FUNCTION_BLOCK UConveyor
VAR
  iStep : INT;
END_VAR
VAR_IN_OUT
  ConveyorIOLeft : ConveyorIO;  (* U的左半边 *)
  ConveyorIORight : ConveyorIO;  (* U的右半边 *)
  ConveyorIODown : ConveyorIO;  (* U的下边一横 *)
  UConveyorIO : UConveyorIO;  (* 顶升,阻挡 *)
END_VAR
VAR
  m_xInitial : BOOL;
  m_tonCylinderOvertime : TON;  (* 气缸超时报警定时器 *)
  m_tCylinderOvertimeCurrent : TIME;
  m_tonExitBarDelay : TON;  (* 退出阻挡器延时 *)
  m_tExitBarDelay : TIME;
  m_xExitBarDelay : BOOL;
  m_TonStep0 : TON;  (* Step为0延时 *)
  m_xStep0 : BOOL;  (* Step为0延时 *)
  m_tStep0 : TIME;  (* Step为0延时 *)
END_VAR
(*                                                                                                          
初始化中增加气缸复位，气缸位置有BUG
//*)
IF NOT m_xInitial THEN
	UConveyorIO.tSetOvertime:=T#5s;
	UConveyorIO.xExitEnable1:=1;
	UConveyorIO.xExitEnable2:=1;
	UConveyorIO.xExitEnable3:=1;
	m_xInitial:=1;
END_IF;
(*外部不用写ConveyorDown的开关，会自己根据来料的产品信息判断停哪个光电*)
IF UConveyorIO.iTask=1 AND ConveyorIODown.diDesConveyorIn=ConveyorIOLeft.diDeviceID THEN
	ConveyorIODown.xCWPresent:=ConveyorIOLeft.xCCWPresent;
ELSIF UConveyorIO.iTask=1 AND ConveyorIODown.diDesConveyorIn=ConveyorIORight.diDeviceID THEN
	ConveyorIODown.xCWPresent:=ConveyorIORight.xCCWPresent;
ELSE
	ConveyorIODown.xCWPresent:=ConveyorIOLeft.xCCWPresent OR ConveyorIORight.xCCWPresent;
END_IF;
(*这里判断什么时候直接放行，左右都不需要，也不是0，就放走*)
IF  NOT(ConveyorIODown.diDesConveyor=ConveyorIOLeft.diDeviceID 
		OR  ConveyorIODown.diDesConveyor=ConveyorIORight.diDeviceID 
		OR ConveyorIODown.diDesConveyor=0) THEN
	UConveyorIO.xPassEnable:=1;
ELSE
	UConveyorIO.xPassEnable:=0;
END_IF;	
IF g_xAuto THEN	
(*	//加个Step为0的延时，防止扫描周期的影响*)
	m_TonStep0(IN:= iStep=0 ,PT:= t#100ms ,Q:= m_xStep0 ,ET:= m_tStep0 );
	(*//这个是留给阻挡动作的时间*)
	m_tonExitBarDelay(IN:=iStep=4 ,PT:= T#1s ,Q:= m_xExitBarDelay ,ET:= m_tExitBarDelay);
CASE UConveyorIO.iTask OF(*这个Task做抢占，可做LastTask保护*)
0:(*各种初始化，能自动去3*)
	ConveyorIODown.xLoad:=0;
	ConveyorIOleft.xLoad:=0;
	ConveyorIORight.xLoad:=0;
	ConveyorIODown.xUnload:=0;
	ConveyorIOLeft.xUnload:=0;
	ConveyorIORight.xUnload:=0;
	ConveyorIODown.xPutInto:=0;
	ConveyorIOLeft.xPutInto:=0;
	ConveyorIORight.xPutInto:=0;	
	UConveyorIO.xExitBarCylinderRetract1:=0;
	UConveyorIO.xExitBarCylinderRetract2:=0;	
	UConveyorIO.xLiftCylinderRetract1:=1;
	UConveyorIO.xLiftCylinderRetract2:=1;
	UConveyorIO.xLiftCylinderExtend1:=0;
	UConveyorIO.xLiftCylinderExtend2:=0;
1:(*上料*)
	CASE iStep OF
	0:(*各种初始化，能自动去3*)
		ConveyorIODown.xLoad:=0;
		ConveyorIOleft.xLoad:=0;
		ConveyorIORight.xLoad:=0;
		ConveyorIODown.xUnload:=0;
		ConveyorIOLeft.xUnload:=0;
		ConveyorIORight.xUnload:=0;
		UConveyorIO.xExitBarCylinderRetract1:=0;
		UConveyorIO.xExitBarCylinderRetract2:=0;
		UConveyorIO.xBatteryError:=0;
		ConveyorIODown.xPutInto:=0;
		ConveyorIOLeft.xPutInto:=0;
		ConveyorIORight.xPutInto:=0;	
	(*	//根据是否有料判断去1还是3，但会等一个延时*)
		IF m_xStep0 AND  ConveyorIODown.xEmpty THEN
			iStep:=1;
		ELSIF m_xStep0 AND NOT ConveyorIODown.xEmpty THEN
			iStep:=3;
		END_IF;	
	1:(*顶升初始化，等load*)
		(*//左顶升*)
		IF UConveyorIO.xLiftCylinderExtendInit1 THEN
			UConveyorIO.xLiftCylinderExtend1:=1;
			UConveyorIO.xLiftCylinderRetract1:=0;
		ELSE
			UConveyorIO.xLiftCylinderExtend1:=0;
			UConveyorIO.xLiftCylinderRetract1:=1;
		END_IF;
	(*	//右顶升*)
		IF UConveyorIO.xLiftCylinderExtendInit2 THEN
			UConveyorIO.xLiftCylinderExtend2:=1;
			UConveyorIO.xLiftCylinderRetract2:=0;
			ELSE
			UConveyorIO.xLiftCylinderExtend2:=0;
			UConveyorIO.xLiftCylinderRetract2:=1;
		END_IF;
		(*//顶升到位，等上料信号*)
		IF 	((UConveyorIO.xLiftCylinderExtendInit1 AND UConveyorIO.xLiftCylinderExtendDetect1)
				OR (NOT UConveyorIO.xLiftCylinderExtendInit1 AND UConveyorIO.xLiftCylinderRetractDetect1))
			AND	((UConveyorIO.xLiftCylinderExtendInit2 AND UConveyorIO.xLiftCylinderExtendDetect2)
		   		OR (NOT UConveyorIO.xLiftCylinderExtendInit2 AND UConveyorIO.xLiftCylinderRetractDetect2))		
			AND	UConveyorIO.xEntryEnable1 THEN(*有上料请求1*)
		   	ConveyorIODown.xLoad:=1;
			iStep:=2;
		END_IF;
	2:(*Load完成*)
		(*去右臂时才需要阻挡1放行,其他情况阻挡1挡住*)
		UConveyorIO.xExitBarCylinderRetract1:=ConveyorIODown.diDesConveyorIn=ConveyorIORight.diDeviceID;
		IF NOT ConveyorIODown.xEmpty THEN
			ConveyorIODown.xLoad:=0;
			ConveyorIOLeft.xPutInto:=1;
			ConveyorIOright.xPutInto:=1;
			istep:=3;
		END_IF;
	3:(*顶升等Unload，这里等有了ExitEnable再顶升，因为可能有地方需要允许了再升降，比如倍速链*)
		(*//电池检测保护，防止把带电池的料框送进去了*)
		IF (ConveyorIODown.diDesConveyor=ConveyorIOLeft.diDeviceID OR ConveyorIODown.diDesConveyor=ConveyorIORight.diDeviceID)
			AND	(UConveyorIO.xBatteryDetect1 OR UConveyorIO.xBatteryDetect2)(*在下面时检测*)
			AND UConveyorIO.xLiftCylinderRetractDetect1 AND UConveyorIO.xLiftCylinderRetractDetect2 THEN
			UConveyorIO.xBatteryError:=1;
		END_IF;	
		(*//左侧顶升控制*)
		IF (ConveyorIODown.diDesConveyor=ConveyorIOLeft.diDeviceID AND UConveyorIO.xExitEnable2 AND NOT UConveyorIO.xBatteryError)THEN
			IF UConveyorIO.xLiftCylinderExtendInit1 THEN
				UConveyorIO.xLiftCylinderExtend1:=0;
				UConveyorIO.xLiftCylinderRetract1:=1;
			ELSE
				UConveyorIO.xLiftCylinderExtend1:=1;
				UConveyorIO.xLiftCylinderRetract1:=0;
			END_IF;
			IF(NOT UConveyorIO.xLiftCylinderExtendInit1 AND UConveyorIO.xLiftCylinderExtendDetect1)
				OR (UConveyorIO.xLiftCylinderExtendInit1 AND UConveyorIO.xLiftCylinderRetractDetect1)THEN
				ConveyorIOLeft.xPutInto:=0;
				ConveyorIOright.xPutInto:=0;
				iStep:=4;
			END_IF;
		END_IF;	
		(*//右侧顶升控制*)
		IF (ConveyorIODown.diDesConveyor=ConveyorIORight.diDeviceID AND UConveyorIO.xExitEnable3 AND NOT UConveyorIO.xBatteryError)THEN
			IF UConveyorIO.xLiftCylinderExtendInit2 THEN
				UConveyorIO.xLiftCylinderExtend2:=0;
				UConveyorIO.xLiftCylinderRetract2:=1;
			ELSE
				UConveyorIO.xLiftCylinderExtend2:=1;
				UConveyorIO.xLiftCylinderRetract2:=0;
			END_IF;
			IF(NOT UConveyorIO.xLiftCylinderExtendInit2 AND UConveyorIO.xLiftCylinderExtendDetect2)
				OR (UConveyorIO.xLiftCylinderExtendInit2 AND UConveyorIO.xLiftCylinderRetractDetect2) THEN
				ConveyorIOLeft.xPutInto:=0;
				ConveyorIOright.xPutInto:=0;
				iStep:=4;
			END_IF;
		END_IF;	
	(*	//直接放行控制*)
		IF UConveyorIO.xPassEnable AND UConveyorIO.xExitEnable1 AND NOT UConveyorIO.xBatteryError THEN
			IF UConveyorIO.xLiftCylinderExtendInit1 THEN
				UConveyorIO.xLiftCylinderExtend1:=1;
				UConveyorIO.xLiftCylinderRetract1:=0;
			ELSE
				UConveyorIO.xLiftCylinderExtend1:=0;
				UConveyorIO.xLiftCylinderRetract1:=1;
			END_IF;
			IF UConveyorIO.xLiftCylinderExtendInit2 THEN
				UConveyorIO.xLiftCylinderExtend2:=1;
				UConveyorIO.xLiftCylinderRetract2:=0;
			ELSE
				UConveyorIO.xLiftCylinderExtend2:=0;
				UConveyorIO.xLiftCylinderRetract2:=1;
			END_IF;
			IF((UConveyorIO.xLiftCylinderExtendInit1 AND UConveyorIO.xLiftCylinderExtendDetect1)
 OR (NOT UConveyorIO.xLiftCylinderExtendInit1 AND UConveyorIO.xLiftCylinderRetractDetect1))
				AND((UConveyorIO.xLiftCylinderExtendInit2 AND UConveyorIO.xLiftCylinderExtendDetect2)
 OR (NOT UConveyorIO.xLiftCylinderExtendInit2 AND UConveyorIO.xLiftCylinderRetractDetect2))THEN
				UConveyorIO.xExitBarCylinderRetract1:=1;
				UConveyorIO.xExitBarCylinderRetract2:=1;
				ConveyorIOLeft.xPutInto:=0;
				ConveyorIOright.xPutInto:=0;
				iStep:=4;
			END_IF;	
		END_IF;
	4:(*Unload完成，回0*)
			IF ConveyorIODown.diDesConveyor=ConveyorIOLeft.diDeviceID AND UConveyorIO.xExitEnable2 AND m_xExitBarDelay THEN
				ConveyorIOLeft.xUnload:=1;
			ELSIF ConveyorIODown.diDesConveyor=ConveyorIORight.diDeviceID AND UConveyorIO.xExitEnable3 AND m_xExitBarDelay THEN
				ConveyorIORight.xUnload:=1;
			ELSIF UConveyorIO.xPassEnable AND UConveyorIO.xExitEnable1 AND m_xExitBarDelay THEN
				ConveyorIODown.xUnload:=1;
			ELSE
				ConveyorIODown.xUnload:=0;
				ConveyorIOLeft.xUnload:=0;
				ConveyorIORight.xUnload:=0;
			END_IF;	
		IF ( (ConveyorIODown.diDesConveyor=ConveyorIOLeft.diDeviceID  AND LDF(TRUE,UConveyorIO.xExitEnable2))
		  OR(ConveyorIODown.diDesConveyor=ConveyorIORight.diDeviceID AND LDF(TRUE,UConveyorIO.xExitEnable3))
		  OR(UConveyorIO.xPassEnable AND LDF(TRUE,UConveyorIO.xExitEnable1)) )AND m_xExitBarDelay  THEN
			ConveyorIODown.xUnload:=0;
			ConveyorIOLeft.xUnload:=0;
			ConveyorIORight.xUnload:=0;
			ConveyorIODown.xPutInto:=1;
			ConveyorIOLeft.xPutInto:=1;
			ConveyorIORight.xPutInto:=1;
			UConveyorIO.xExitBarCylinderRetract1:=0;
			UConveyorIO.xExitBarCylinderRetract2:=0;
			iStep:=0;
		END_IF;
	END_CASE;
2:(*左下料*)
	CASE iStep OF
	0:(*各种初始化，能自动去3*)
		ConveyorIODown.xLoad:=0;
		ConveyorIOleft.xLoad:=0;
		ConveyorIORight.xLoad:=0;
		ConveyorIODown.xUnload:=0;
		ConveyorIOLeft.xUnload:=0;
		ConveyorIORight.xUnload:=0;
		UConveyorIO.xBatteryError:=0;
		UConveyorIO.xExitBarCylinderRetract1:=0;
		UConveyorIO.xExitBarCylinderRetract2:=0;
		ConveyorIODown.xPutInto:=0;
		ConveyorIOLeft.xPutInto:=0;
		ConveyorIORight.xPutInto:=0;
		IF m_xStep0 AND  ConveyorIODown.xEmpty THEN
			iStep:=1;
		ELSIF m_xStep0 AND NOT ConveyorIODown.xEmpty THEN
			iStep:=3;
		END_IF;	
	1:(*左顶升动作，等load*)
		IF UConveyorIO.xLiftCylinderExtendInit1 THEN
			UConveyorIO.xLiftCylinderExtend1:=0;
			UConveyorIO.xLiftCylinderRetract1:=1;
			ELSE
			UConveyorIO.xLiftCylinderExtend1:=1;
			UConveyorIO.xLiftCylinderRetract1:=0;
		END_IF;
		IF ((NOT UConveyorIO.xLiftCylinderExtendInit1 AND UConveyorIO.xLiftCylinderExtendDetect1)
			OR ( UConveyorIO.xLiftCylinderExtendInit1 AND UConveyorIO.xLiftCylinderRetractDetect1))
			AND UConveyorIO.xEntryEnable2 THEN(*有上料请求1*)
		   	ConveyorIOLeft.xLoad:=1;
			iStep:=2;
		END_IF;
	2:(*Load完成*)
		IF NOT ConveyorIOLeft.xEmpty THEN
			ConveyorIOLeft.xLoad:=0;
			ConveyorIODown.xPutInto:=1;
			ConveyorIODown.diDesConveyor:=ConveyorIOLeft.diDesConveyor;
			istep:=3;
		END_IF;
	3:(*顶升等Unload，这里等有了ExitEnable再顶升，因为可能有地方需要允许了再升降，比如倍速链*)
		UConveyorIO.xExitBarCylinderRetract1:=1;
		UConveyorIO.xExitBarCylinderRetract2:=1;
		IF  UConveyorIO.xExitEnable1 THEN
			IF UConveyorIO.xLiftCylinderExtendInit1 THEN
				UConveyorIO.xLiftCylinderExtend1:=1;
				UConveyorIO.xLiftCylinderRetract1:=0;
			ELSE
				UConveyorIO.xLiftCylinderExtend1:=0;
				UConveyorIO.xLiftCylinderRetract1:=1;
			END_IF;
			IF(( UConveyorIO.xLiftCylinderExtendInit1 AND UConveyorIO.xLiftCylinderExtendDetect1)
				OR (NOT UConveyorIO.xLiftCylinderExtendInit1 AND UConveyorIO.xLiftCylinderRetractDetect1))THEN
				ConveyorIODown.xPutInto:=0;
				iStep:=4;
			END_IF;	
		END_IF;
	4:(*Unload完成，回0*)
		IF  UConveyorIO.xExitEnable1 AND m_xExitBarDelay THEN
			ConveyorIODown.xUnload:=1;
		ELSE
			ConveyorIODown.xUnload:=0;
		END_IF;	
		IF NOT UConveyorIO.xExitEnable1 AND m_xExitBarDelay   THEN
			ConveyorIODown.xUnload:=0;
			ConveyorIOLeft.xUnload:=0;
			ConveyorIORight.xUnload:=0;
			ConveyorIODown.xPutInto:=1;
			ConveyorIOLeft.xPutInto:=1;
			ConveyorIORight.xPutInto:=1;
			UConveyorIO.xExitBarCylinderRetract1:=0;
			UConveyorIO.xExitBarCylinderRetract2:=0;
			iStep:=0;
		END_IF;
	END_CASE;
3:(*上料到出口*)
	CASE iStep OF
	0:(*各种初始化，能自动去3*)
		ConveyorIODown.xLoad:=0;
		ConveyorIOleft.xLoad:=0;
		ConveyorIORight.xLoad:=0;
		ConveyorIODown.xUnload:=0;
		ConveyorIOLeft.xUnload:=0;
		ConveyorIORight.xUnload:=0;
		UConveyorIO.xBatteryError:=0;
		UConveyorIO.xExitBarCylinderRetract1:=0;
		UConveyorIO.xExitBarCylinderRetract2:=0;
		ConveyorIODown.xPutInto:=0;
		ConveyorIOLeft.xPutInto:=0;
		ConveyorIORight.xPutInto:=0;
		IF m_xStep0 AND  ConveyorIODown.xEmpty THEN
			iStep:=1;
		ELSIF m_xStep0 AND NOT ConveyorIODown.xEmpty THEN
			iStep:=3;
		END_IF;	
	1:(*右顶升动作，等load*)
		IF UConveyorIO.xLiftCylinderExtendInit2 THEN
			UConveyorIO.xLiftCylinderExtend2:=0;
			UConveyorIO.xLiftCylinderRetract2:=1;
		ELSE
			UConveyorIO.xLiftCylinderExtend2:=1;
			UConveyorIO.xLiftCylinderRetract2:=0;
		END_IF;
		IF ((NOT UConveyorIO.xLiftCylinderExtendInit2 AND UConveyorIO.xLiftCylinderExtendDetect2)
			OR ( UConveyorIO.xLiftCylinderExtendInit2 AND UConveyorIO.xLiftCylinderRetractDetect2))
			AND UConveyorIO.xEntryEnable3 THEN(*有上料请求1*)
		   	ConveyorIORight.xLoad:=1;
			iStep:=2;
		END_IF;
	2:(*Load完成*)
		IF NOT ConveyorIORight.xEmpty THEN
			ConveyorIORight.xLoad:=0;
			ConveyorIODown.diDesConveyor:=ConveyorIORight.diDesConveyor;
			ConveyorIODown.xPutInto:=1;
			istep:=3;
		END_IF;
	3:(*顶升恢复等Unload，这里等有了ExitEnable再顶升，因为可能有地方需要允许了再升降，比如倍速链*)
		UConveyorIO.xExitBarCylinderRetract2:=1;
		IF  UConveyorIO.xExitEnable1 THEN(**)
			IF UConveyorIO.xLiftCylinderExtendInit2 THEN
				UConveyorIO.xLiftCylinderExtend2:=1;
				UConveyorIO.xLiftCylinderRetract2:=0;
			ELSE
				UConveyorIO.xLiftCylinderExtend2:=0;
				UConveyorIO.xLiftCylinderRetract2:=1;
			END_IF;
		END_IF;
		IF UConveyorIO.xExitEnable1 THEN(**)
			IF(( UConveyorIO.xLiftCylinderExtendInit2 AND UConveyorIO.xLiftCylinderExtendDetect2)
				OR (NOT UConveyorIO.xLiftCylinderExtendInit2 AND UConveyorIO.xLiftCylinderRetractDetect2))THEN
				ConveyorIODown.xPutInto:=0;
				iStep:=4;
			END_IF;	
		END_IF;
	4:(*Unload完成，回0*)
		IF  UConveyorIO.xExitEnable1 AND m_xExitBarDelay THEN
			ConveyorIODown.xUnload:=1;
		ELSE
			ConveyorIODown.xUnload:=0;
		END_IF;	
		IF NOT UConveyorIO.xExitEnable1 AND m_xExitBarDelay  THEN
			ConveyorIODown.xUnload:=0;
			ConveyorIOLeft.xUnload:=0;
			ConveyorIORight.xUnload:=0;
			ConveyorIODown.xPutInto:=1;
			ConveyorIOLeft.xPutInto:=1;
			ConveyorIORight.xPutInto:=1;
			UConveyorIO.xExitBarCylinderRetract1:=0;
			UConveyorIO.xExitBarCylinderRetract2:=0;
			iStep:=0;
		END_IF;
	END_CASE;
END_CASE;(*iTask*)
END_IF;(*g_xAuto那个IF*)
(*复位程序*)
IF (g_xResetSingle AND  (g_diDeviceIDSelect=ConveyorIOLeft.diDeviceID 
 	 OR g_diDeviceIDSelect=ConveyorIORight.diDeviceID
 	 OR g_diDeviceIDSelect=ConveyorIODown.diDeviceID))
	OR LDP(TRUE,UConveyorIO.xLiftCylinderExtendInit1) 
	OR LDF(TRUE,UConveyorIO.xLiftCylinderExtendInit1) 
	OR LDP(TRUE,UConveyorIO.xPutInto)  THEN
	ConveyorIODown.xPutInto:=1;
	ConveyorIOLeft.xPutInto:=1;
	ConveyorIORight.xPutInto:=1;
	iStep:=0;
END_IF;
(*手动*)
IF g_xManual  THEN
	iStep:=0;
	ConveyorIODown.xLoad:=0;
	ConveyorIOleft.xLoad:=0;
	ConveyorIORight.xLoad:=0;
	ConveyorIODown.xUnload:=0;
	ConveyorIOLeft.xUnload:=0;
	ConveyorIORight.xUnload:=0;
	ConveyorIODown.xPutInto:=0;
	ConveyorIOLeft.xPutInto:=0;
	ConveyorIORight.xPutInto:=0;
	UConveyorIO.xBatteryError:=0;
	UConveyorIO.xLiftCylinderExtend1:=UConveyorIO.xLiftCylinderExtendButton1 AND NOT UConveyorIO.xLiftCylinderRetractButton1;
	UConveyorIO.xLiftCylinderRetract1:=UConveyorIO.xLiftCylinderRetractButton1 AND NOT UConveyorIO.xLiftCylinderExtendButton1;
	UConveyorIO.xLiftCylinderExtend2:=UConveyorIO.xLiftCylinderExtendButton2 AND NOT UConveyorIO.xLiftCylinderRetractButton2;
	UConveyorIO.xLiftCylinderRetract2:=UConveyorIO.xLiftCylinderRetractButton2 AND NOT UConveyorIO.xLiftCylinderExtendButton2;
	UConveyorIO.xExitBarCylinderRetract1:=UConveyorIO.xExitBarCylinderRetractButton1;
	UConveyorIO.xExitBarCylinderRetract2:=UConveyorIO.xExitBarCylinderRetractButton2;
END_IF;	
(*气缸超时报警*)
m_tonCylinderOvertime(IN:= (UConveyorIO.xLiftCylinderExtend1 AND NOT UConveyorIO.xLiftCylinderExtendDetect1) 
 		OR  (UConveyorIO.xLiftCylinderRetract1 AND NOT UConveyorIO.xLiftCylinderRetractDetect1)
 		OR	(UConveyorIO.xLiftCylinderExtend2 AND NOT UConveyorIO.xLiftCylinderExtendDetect2) 
 		OR  (UConveyorIO.xLiftCylinderRetract2 AND NOT UConveyorIO.xLiftCylinderRetractDetect2),
 PT:= UConveyorIO.tSetOvertime ,Q:=UConveyorIO.xOvertimeAlarm ,ET:=m_tCylinderOvertimeCurrent );
END_FUNCTION_BLOCK

PROGRAM 批量复制专用

END_PROGRAM

FUNCTION_BLOCK FanucRobot
VAR_IN_OUT
  FanucRobotIO : FanucRobotIO;
END_VAR
VAR
  m_iSNO : INT;
  m_xPNSPass : BOOL;  (* 收到程序号 *)
  m_tonStartDelay : TON;  (* 启动延时 *)
  m_xStartDelay : BOOL;
  m_tStartDelayCurrentTime : TIME;
END_VAR
(***********************************************************
发那科机器人自动启动程序


***********************************************************)

(*无自动状态，示教盒处于本地状态，把各标志位复位*)
IF FanucRobotIO.i_xTPENBL AND NOT g_xAuto THEN
	FanucRobotIO.o_xPNSTROBE:=0;
	FanucRobotIO.o_xCSTOPI:=0;
	FanucRobotIO.o_xPROD_START:=0;
	FanucRobotIO.o_xRESET:=0;
END_IF;
(*远程模式*)
IF g_xAuto THEN
	FanucRobotIO.o_xREMOTE:=1;
	ELSE
	FanucRobotIO.o_xREMOTE:=0;
END_IF;
(*程序启动后复位启动标志位*)
IF FanucRobotIO.i_xPROG_RUN AND FanucRobotIO.i_xBUSY THEN
	FanucRobotIO.i_xCommandStart:=0;
END_IF;
(*示教盒旋清除报警*)
IF ldf(TRUE,FanucRobotIO.i_xTPENBL)THEN
	FanucRobotIO.o_xRESET:=1;
	FanucRobotIO.o_xCSTOPI:=1;
END_IF;
(*启动程序号条件*)
IF FanucRobotIO.i_xSYSRDY 
	AND FanucRobotIO.i_xCMDENBL
	AND FanucRobotIO.i_xCommandStart
	AND NOT FanucRobotIO.i_xPROG_RUN 
	AND NOT FanucRobotIO.i_xBUSY THEN
	FanucRobotIO.o_xRESET:=0;
	FanucRobotIO.o_xCSTOPI:=0;
	IF FanucRobotIO.i_iMotionNumber <> 0 (*只要动作编号不为0，就给他信号*)
		AND NOT FanucRobotIO.o_xPNSTROBE THEN
		FanucRobotIO.o_xPNSTROBE:=1;
		FanucRobotIO.o_xPROD_START:=1;
		FanucRobotIO.o_iPNS:=FanucRobotIO.i_iMotionNumber;(*并把任务号传给他*)
	END_IF;
	(*程序号校验*)
	IF FanucRobotIO.i_xSNACK THEN(*数据传回之后再校验*)
		m_iSNO:=BITARR_TO_INT(FanucRobotIO.i_arrxSNO[0] , 8 );
		IF m_iSNO=FanucRobotIO.o_iPNS THEN
			m_xPNSPass:=1;(*校验成功,等100MS复位Start信号*)
			FanucRobotIO.o_xPNSTROBE:=0;
		ELSE
			FanucRobotIO.o_xPNSFailed:=1;(*校验失败*)
			FanucRobotIO.o_xPROD_START:=0;(*立刻复位，不生成任务*)
		END_IF;
	END_IF;
END_IF;
m_tonStartDelay(IN:= m_xPNSPass ,PT:= T#100ms ,Q:= m_xStartDelay ,ET:=m_tStartDelayCurrentTime );
IF m_xStartDelay THEN
	FanucRobotIO.o_xPROD_START:=0;
	FanucRobotIO.i_xCommandStart:=0;
	m_xPNSPass:=0;
END_IF;
END_FUNCTION_BLOCK

FUNCTION_BLOCK ConveyorCommunication
VAR_IN_OUT
  ConveyorIO : ConveyorIO;
  CommunicationIO : CommunicationIO;
END_VAR
VAR_OUTPUT
  o_iErrorNub : INT;  (* 错误代码 *)
END_VAR
VAR
  o_xReqSuccess : BOOL;  (* 请求成功 *)
END_VAR
(********************************************************************************)
(*
DB1区(PC->PLC)15个字		
"字(16位）序号
(从1开始)"			功能描述  	具体参数解释
1 请求确认	"  1：复位
				   				2：读码(入库申请）成功
				   				3：取放货完成 
   			4：旋转
   			5：不旋转
   			101：条码空
   			102：条码规则校验失败
   			103：步号校验失败
   			104：无库位可用 
"
2	预留	
3	预留	
4	预留	
5	预留	
6	读写标志位	"  				1：写入数据
   			2：读数据完成"
7	任务处理标志	"  				１：复位
   			２：完成"
8	命令字	"
   			21-送出（任务起点与终点不同，即向下一台输送机移载）
   			22：叠盘
"
9	任务号	"   1~65535唯一任务标识"
10	目标设备号   只有送出任务才有效
11		
12	筐码后4位	
				

DB2区(PLC->PC)15个字			
"字(16位）序号
(从1开始)"	功能描述	具体参数解释	
1	请求状态	"１：复位
２：请求"	实时状态，没有时序交互
2	强制入库(预留）	"１：复位
２：强制入库"	
3	预留(叠盘数量）	只对叠盘工位有效	
4	预留		
5			
6	读写标志位	"1：写入数据
2：读数据完成"	"有交互
时序"
7	设备状态	"1:空闲
2：工作中
3:任务完成（只有目标设备才会报任务完成）
４：故障"	
8	任务号	1~65535唯一任务标识，当输送任务执行完成后，将PC下发的任务号上报	
9	筐码后4位		
10	预留		
11			
			





2018.8.3 YAO 1.0
*)
(********************************************************************************)
(*//请求状态*)
IF ConveyorIO.xEmpty THEN
	CommunicationIO.o_iRequestPLCPC:=1;
	ELSE
	CommunicationIO.o_iRequestPLCPC:=2;
END_IF;
(*//请求确认*)
CASE CommunicationIO.i_iResponsPCPLC OF 
	0:;
	1:;(*//复位*)
	2:(*//读码（入库申请）成功*)
	o_xReqSuccess:=1;
	3:(*//取放货完成*)
	ConveyorIO.xPutInto:=1; 
	4:(*//旋转*)
	;
	5:(*//不旋转*)
	;
	101:(*//条码空*)
	o_iErrorNub:=101;
	102:(*//条码规则检验失败*)
	o_iErrorNub:=102;
	103:(*//步号校验失败*)
	o_iErrorNub:=103;
	104:(*//无库位可用*)
	o_iErrorNub:=104;
END_CASE;
IF CommunicationIO.i_iResponsPCPLC <> 3 THEN
	ConveyorIO.xPutInto:=0;
END_IF;
IF CommunicationIO.i_iResponsPCPLC <> 2 THEN
	o_xReqSuccess:=0;
END_IF;
IF CommunicationIO.i_iResponsPCPLC < 100 THEN
	o_iErrorNub:=0;
END_IF;

(*//读写标志位写入数据*)
IF LDP(TRUE,CommunicationIO.i_iReadWriteFlagPCPLC = 1) THEN
	ConveyorIO.iTaskID := CommunicationIO.i_iTaskIDPCPLC;
	ConveyorIO.diDesConveyor := CommunicationIO.i_diDestinationDevicePCPLC;
	ConveyorIO.iProductCategory := CommunicationIO.i_iProductIDPCPLC;
END_IF;
(*//数据校验，并返回握手信号*)
IF CommunicationIO.i_iReadWriteFlagPCPLC = 1 
	AND ConveyorIO.iTaskID<>0
	AND ConveyorIO.diDesConveyor<>0 
	AND ConveyorIO.iProductCategory<>0 
	THEN
	CommunicationIO.o_iReadWriteFlagPLCPC:=2;
	ELSE
	CommunicationIO.o_iReadWriteFlagPLCPC:=1;
END_IF;
(*//数据校验*)
IF CommunicationIO.i_iReadWriteFlagPCPLC = 1 
	AND (ConveyorIO.iTaskID<>0
	OR ConveyorIO.diDesConveyor<>0 
	OR ConveyorIO.iProductCategory<>0) 
	THEN
	o_iErrorNub:=50;(*//任务数据不完整*)
END_IF;
(*//设备状态*)
IF ConveyorIO.diDesConveyor = ConveyorIO.diDeviceID AND NOT ConveyorIO.xEmpty THEN(*//目标地址=当前地址*)
	CommunicationIO.o_iDeviceStatusPLCPC:=3;(*//任务完成*)
	CommunicationIO.o_iProductIDPLCPC:=ConveyorIO.iProductCategory;(*//条码号上传*)
	CommunicationIO.o_iTaskIDPLCPC:=ConveyorIO.iTaskID;(*//任务号上传*)
	ELSIF ConveyorIO.xBusy THEN
	CommunicationIO.o_iDeviceStatusPLCPC:=2;(*//工作中*)
	ELSIF ConveyorIO.xError THEN
	CommunicationIO.o_iDeviceStatusPLCPC:=4;(*//故障*)
	ELSE
	CommunicationIO.o_iDeviceStatusPLCPC:=1;(*//空闲*)
	CommunicationIO.o_iProductIDPLCPC:=0;(*//条码号复位*)
	CommunicationIO.o_iTaskIDPLCPC:=0;(*//任务号复位*)
END_IF;
END_FUNCTION_BLOCK

FUNCTION_BLOCK PackCommunication
VAR_IN_OUT
  ConveyorIO : ConveyorIO;
  PackCommunicationIO : PackCommunicationIO;
  FanucRobotIO : FanucRobotIO;
END_VAR
VAR_OUTPUT
  o_iErrorNub : INT;
  o_xReqSuccess : BOOL;
END_VAR
VAR
  m_xReqSuccess : BOOL;
  m_iStep : INT;
  m_arrwCode : ARRAY [1..8] OF BatteryCode;
END_VAR
VAR_INPUT
  i_arrxPresentDetect : ARRAY [1..8] OF BOOL;
END_VAR
VAR
  m_iCoordinateX : INT;
  m_iCoordinateY : INT;
  m_arriPresentDetect : ARRAY [1..8] OF INT;
  ii : INT;
END_VAR
VAR CONSTANT
  MAX_ROW : INT := 8;
  MAX_COLUMN : INT := 8;
END_VAR
VAR
  m_xSupplement : BOOL;
END_VAR
VAR CONSTANT
  ROW_TIMES : INT := 1;
  GET_QUANTITY : INT := 8;
END_VAR
VAR
  m_iRowReminder : INT;
  m_xEno : BOOL;
  m_iRowReminderTemp : INT;
END_VAR
(***************************************************************************)
(*
DB1区(PC->PLC)10个字		
"字(16位）序号
(从1开始)"	功能描述	具体参数解释
1	请求确认	"1：复位
2：读码(入库申请）成功
101：条码空
102：条码规则校验失败
103：步号校验失败
"
2	放行	"1：复位
2：完成,放行
3：撤销完成 "
3	单次装载应答	"1：复位
2：允许开始"
4	单次装载处理完成	"1：复位
2：完成
3：电芯为空"
)*
DB2区(PLC->PC)200个字		
"字(16位）序号
(从1开始)"	功能描述	具体参数解释
1	装载请求	"１：复位
２：请求"
2	装载全部完成	"1：复位
2：请求 "
3	单次装载请求	"1：复位
2：请求 "
4	单次装载完成	"1：复位
2：完成"
5	行坐标	从1开始
6	列坐标	从1开始
7	电芯码(15*11=165)	"电芯码24字符，
占12个字，加上预留的每个分配15个字"

顺序执行步骤
0  初始化
1  框码扫码请求
2  单次抓取请求
3  整排抓取
4  补料
5  完成


(***************************************************************************)
m_iRowReminder:= ( m_iCoordinateX-1 MOD GET_QUANTITY )+1;(*//通过位置与抓取数量取余数，判断是否的抓取位置为一排的最后一个*)
CASE m_iStep OF
	0:;(*//初始化*)
	m_iStep:=1;
	1:(*发送框码的扫码请求*)
	IF NOT ConveyorIO.xEmpty AND NOT FanucRobotIO.io_xMutexLock THEN
		PackCommunicationIO.o_iRequestPLCPC:=2;
		ELSE
		PackCommunicationIO.o_iRequestPLCPC:=1;
	END_IF;
	(*//请求确认*)
	CASE PackCommunicationIO.i_iResponsPCPLC OF 
		0:;
		1:;(*//复位*)
		2:(*//读码（入库申请）成功*)
		m_iStep:=2;
		m_xSupplement:=0;
		m_iCoordinateX:=1;(*//框码扫码成功后把坐标改为1,1*)
		m_iCoordinateY:=1;
		FanucRobotIO.io_xMutexLock:=1;
		3:(*//取放货完成*)
		ConveyorIO.xPutInto:=1; 
		4:(*//旋转*)
		;
		5:(*//不旋转*)
		;
		101:(*//条码空*)
		o_iErrorNub:=101;
		m_iStep:=0;
		102:(*//条码规则检验失败*)
		o_iErrorNub:=102;
		m_iStep:=0;
		103:(*//步号校验失败*)
		o_iErrorNub:=103;
		m_iStep:=0;
		104:(*//无库位可用*)
		o_iErrorNub:=104;
		m_iStep:=0;
	END_CASE;
	2:(*//单次抓取请求，分为单次多个产品抓取与补料程序*)
	IF FanucRobotIO.i_xSYSRDY 
		AND NOT FanucRobotIO.i_xBUSY
		AND NOT FanucRobotIO.i_xPROG_RUN
		AND i_arrxPresentDetect[1] 
		AND PackCommunicationIO.i_iSinglePackResponsePCPLC=1 THEN(*//机器人准备就绪、组装下线有料*)
		PackCommunicationIO.o_iSinglePackRequestPLCPC:=2;
	END_IF;
	IF (*LDP(TRUE,PackCommunicationIO.i_iSinglePackResponsePCPLC=2)*) PackCommunicationIO.i_iSinglePackResponsePCPLC=2 THEN(*//请求成功*)
		PackCommunicationIO.o_iSinglePackRequestPLCPC:=1;(*//复位请求*)
		IF m_xSupplement THEN(*//补料标志位，为1进行补料操作，为0进行整排抓取*)
			m_iStep:=4;(*//补料*)
			ELSE
		 	m_iStep:=3;(*//整排抓取*)
			FOR ii:=1 TO GET_QUANTITY BY 1 DO(*//记录哪个位置缺料*)
				IF i_arrxPresentDetect[ii] THEN(*//传感器检测*)
 m_arriPresentDetect[ii]:=0;
 ELSE
 m_arriPresentDetect[ii]:=ii;(*//记录缺料的位置*)
				END_IF;
			END_FOR;
		END_IF;
	END_IF;
	3:  (*//整排抓取*)
	FanucRobotIO.o_iPNS:=10101;(*//步骤号*)
	FanucRobotIO.o_uiOffset_X:=m_iCoordinateX;
	FanucRobotIO.o_uiOffset_Y:=m_iCoordinateY;
	PackCommunicationIO.o_iXCoordinatePLCPC:=m_iCoordinateX;(*//放置位置发送给上位机*)
	PackCommunicationIO.o_iYCoordinatePLCPC:=m_iCoordinateY;	
	IF LDF(TRUE,FanucRobotIO.i_xBUSY OR FanucRobotIO.i_xPROG_RUN) THEN(*//抓取动作完成*)
		FOR ii:=1 TO GET_QUANTITY BY 1 DO (*//判断有无补料信息*)
			IF m_arriPresentDetect[ii]<>0  THEN(*//有补料*)(*//补料不是最后一个的算法*)
				m_iCoordinateX:=m_arriPresentDetect[ii]+((m_iCoordinateX-1)/GET_QUANTITY)*GET_QUANTITY;
				m_xSupplement:=1;
				m_iStep:=2;(*//有补料*)
				EXIT;
			END_IF;			
		END_FOR;
		IF ii=GET_QUANTITY+1  THEN  (*//无补料*)
			m_xSupplement:=0;
			IF m_iCoordinateY = MAX_ROW (*//达到最大列*)
				AND ((m_iCoordinateX-1)/GET_QUANTITY+1=ROW_TIMES) 
				THEN(*//偏移量为最大的值时,排抓取为最后一排*)
				m_iStep:=5;(*//装盘完成*)
				ELSE
				m_iStep:=2;(*//请求下一次装盘*)			
				IF (m_iCoordinateX-1)/GET_QUANTITY+1=ROW_TIMES THEN
 m_iCoordinateX:=1;                                              (*//开始执行下一列*)
 m_iCoordinateY:=m_iCoordinateY+1;
 ELSE
 m_iCoordinateX:=((m_iCoordinateX-1)/GET_QUANTITY+1)*GET_QUANTITY+1;
				END_IF;
			END_IF;
		END_IF;
	END_IF;
	4: (*//补料*)
	FanucRobotIO.o_iPNS:=10102;(*//步骤号*)
	FanucRobotIO.o_uiOffset_X:=m_iCoordinateX;
	FanucRobotIO.o_uiOffset_Y:=m_iCoordinateY;
	PackCommunicationIO.o_iXCoordinatePLCPC:=m_iCoordinateX;(*//放置位置发送给上位机*)
	PackCommunicationIO.o_iYCoordinatePLCPC:=m_iCoordinateY;
	IF LDF(TRUE,FanucRobotIO.i_xBUSY OR FanucRobotIO.i_xPROG_RUN) THEN(*//抓取动作完成*)
		FOR ii:=m_iRowReminder+1 TO GET_QUANTITY BY 1 DO (*//判断有无补料信息*)
			IF m_arriPresentDetect[ii]<>0  THEN(*//有补料*)(*//补料不是最后一个的算法*)
				m_iCoordinateX:=m_arriPresentDetect[ii]+((m_iCoordinateX-1)/GET_QUANTITY)*GET_QUANTITY;
				m_xSupplement:=1;
				m_iStep:=2;(*//有补料*)
				EXIT;
			END_IF;	
		END_FOR;
		IF ii=GET_QUANTITY+1  THEN  (*//无补料*)
			m_xSupplement:=0;
			IF m_iCoordinateY = MAX_ROW (*//达到最大列*)
				AND ((m_iCoordinateX-1)/GET_QUANTITY+1=ROW_TIMES)
				THEN(*//偏移量为最大的值时,排抓取为最后一排*)
				m_iStep:=5;(*//装盘完成*)
				ELSE
				m_iStep:=2;(*//请求下一次装盘*)			
				IF (m_iCoordinateX-1)/GET_QUANTITY+1=ROW_TIMES THEN
 m_iCoordinateX:=1;                                              (*//开始执行下一列*)
 m_iCoordinateY:=m_iCoordinateY+1;
 ELSE
 m_iCoordinateX:=((m_iCoordinateX-1)/GET_QUANTITY+1)*GET_QUANTITY+1;(*//这一列继续往后排*)
				END_IF;
			END_IF;
		END_IF;
	END_IF;
	5: (*//完成*)
	PackCommunicationIO.o_iSinglePackDonePLCPC:=2;
	IF PackCommunicationIO.i_iSinglePackDoneAknPCPLC =2 THEN
		PackCommunicationIO.o_iSinglePackDonePLCPC:=1;
		m_iCoordinateX:=1;
		m_iCoordinateY:=1;
		FanucRobotIO.io_xMutexLock:=0;
	END_IF;
	IF ConveyorIO.xEmpty AND PackCommunicationIO.o_iSinglePackDonePLCPC=1 THEN
		m_iStep:=1;
	END_IF;
END_CASE;
END_FUNCTION_BLOCK

PROGRAM START
IF g_xReset THEN
	SM50:=1;
	ELSE
	SM50:=0;
END_IF;
CASE g_iState OF
	0: (*手动*)
	g_xManual:=1;
	g_xAuto:=0;	
	g_xStackLampAmber:=1;
	g_xStackLampGreen:=0;
	g_xRemoteAuto:=0;
	g_xAutoLamp:=0;
	1:(*自动*)
	g_xManual:=0;
	g_xAuto:=1;
	g_xStackLampGreen:=1;
	g_xStackLampAmber:=0;
	g_xRemoteAuto:=0;
	g_xAutoLamp:=1;
	2:	(*远程自动*)
	g_xRemoteAuto:=1;
	g_xStackLampGreen:=1;
	g_xStackLampAmber:=0;
	g_xAuto:=0;
	g_xManual:=0;
	g_xAutoLamp:=0;
	3:(*自动未启动*)
	g_xRemoteAuto:=1;
	g_xStackLampGreen:=SM412;
	g_xStackLampAmber:=0;
	g_xAuto:=0;
	g_xManual:=0;	
	g_xAutoLamp:=0;
END_CASE;

IF g_xAutoSwitch AND g_xAutoStart  THEN  
	g_iState:=1;
END_IF;

IF g_xAutoSwitch AND (g_iState<>1 OR NOT g_xStop)  THEN  
	g_iState:=3;
END_IF;

g_xStackLampRed:=g_xAlarm AND SM412;
g_xBuzzer:=g_xAlarm AND SM412 AND NOT g_xMute;

IF LDF(TRUE,g_xAlarm) THEN
	g_xMute:=0;
END_IF;

IF NOT g_xAutoSwitch  OR g_xEStop=0 THEN 
	g_iState:=0;
END_IF;
IF g_xRemoteAutoStart THEN
	g_iState:=2;
END_IF;
IF g_xPause AND SM412 THEN
	g_xStackLampGreen:=0;
	g_xStackLampAmber:=0;
END_IF;
END_PROGRAM
